FUNCTION "LKinCtrl_CallMC_Reset_SyncAxis" : Void   // FC35024, SCL
{ S7_Optimized_Access := 'TRUE' }
VERSION : 0.1
   VAR_INPUT
      syncAxisIn : TO_SynchronousAxis;   // SynchronousAxis to access
      execute : Bool;   // execute signal for MC_RESET
      restart : Bool;   // restart signal for MC_RESET
   END_VAR
   VAR_IN_OUT
      instMC_Reset : MC_RESET;   // multi instance of MC_RESET
   END_VAR
BEGIN
   //================================================================================
   // SIEMENS AG
   // (c)Copyright 2019 All Rights Reserved
   //--------------------------------------------------------------------------------
   // Library: LKinCtrl
   // Tested with: S7-1517T-3 PN
   // Engineering: TIA Portal V15
   // Restrictions: -
   // Requirements: S7-1500T FW 2.5
   // Functionality: Call MC_Home
   // Support: tech.team.motioncontrol@siemens.com
   // Note: Parameter comments are only available in language 'English (United States)'
   //-----------------------------------------------------------------------------
   // Change log table:
   // Version    Date          Expert in charge    Changes applied
   // 01.00.00   27.02.2019    JR                  First released version
   //===========================================================================================

   // call MC_Reset
   #instMC_Reset(Axis:=#syncAxisIn,
                 Execute:=#execute,
                 Restart:=#restart);
END_FUNCTION

FUNCTION "LKinCtrl_CallMC_Reset_PosAxis" : Void   // FC35025, SCL
{ S7_Optimized_Access := 'TRUE' }
VERSION : 0.1
   VAR_INPUT
      posAxisIn : TO_PositioningAxis;   // PositioningAxis to access
      execute : Bool;   // execute signal for MC_RESET
      restart : Bool;   // restart signal for MC_RESET
   END_VAR
   VAR_IN_OUT
      instMC_Reset : MC_RESET;   // multi instance of MC_RESET
   END_VAR
BEGIN
   //================================================================================
   // SIEMENS AG
   // (c)Copyright 2019 All Rights Reserved
   //--------------------------------------------------------------------------------
   // Library: LKinCtrl
   // Tested with: S7-1517T-3 PN
   // Engineering: TIA Portal V15
   // Restrictions: -
   // Requirements: S7-1500T FW 2.5
   // Functionality: Call MC_Reset
   // Support: tech.team.motioncontrol@siemens.com
   // Note: Parameter comments are only available in language 'English (United States)'
   //-----------------------------------------------------------------------------
   // Change log table:
   // Version    Date          Expert in charge    Changes applied
   // 01.00.00   27.02.2019    JR                  First released version
   //===========================================================================================

   // call MC_Reset
   #instMC_Reset(Axis:=#posAxisIn,
                 Execute:=#execute,
                 Restart:=#restart);
END_FUNCTION

FUNCTION "LKinCtrl_CallMC_Home_SyncAxis" : Void   // FC35026, SCL
{ S7_Optimized_Access := 'TRUE' }
VERSION : 0.1
   VAR_INPUT
      syncAxisIn : TO_SynchronousAxis;   // SynchronousAxis to access
      execute : Bool;   // execute trigger
      position : LReal;   // home position
      mode : Int;   // homing mode
   END_VAR
   VAR_IN_OUT
      instMC_Home : MC_HOME;   // multi instance MC_HOME
   END_VAR
BEGIN
   //================================================================================
   // SIEMENS AG
   // (c)Copyright 2019 All Rights Reserved
   //--------------------------------------------------------------------------------
   // Library: LKinCtrl
   // Tested with: S7-1517T-3 PN
   // Engineering: TIA Portal V15
   // Restrictions: -
   // Requirements: S7-1500T FW 2.5
   // Functionality: Call MC_Home
   // Support: tech.team.motioncontrol@siemens.com
   // Note: Parameter comments are only available in language 'English (United States)'
   //-----------------------------------------------------------------------------
   // Change log table:
   // Version    Date          Expert in charge    Changes applied
   // 01.00.00   27.02.2019    JR                  First released version
   //===========================================================================================

   // call MC_Home
   #instMC_Home(Axis:=#syncAxisIn,
                Execute:=#execute,
                Position:=#position,
                Mode:=#mode);
END_FUNCTION

FUNCTION "LKinCtrl_CallMC_Power_PosAxis" : Void   // FC35027, SCL
{ S7_Optimized_Access := 'TRUE' }
VERSION : 0.1
   VAR_INPUT
      posAxisIn : TO_PositioningAxis;   // PositioningAxis to access
      enable : Bool;   // execute signal for MC_RESET
      startMode : DInt;   // startMode of axis
      stopMode : Int;   // stopMode of axis
   END_VAR
   VAR_IN_OUT
      instMC_Power : MC_POWER;   // multi instance of MC_RESET
   END_VAR
BEGIN
   //================================================================================
   // SIEMENS AG
   // (c)Copyright 2019 All Rights Reserved
   //--------------------------------------------------------------------------------
   // Library: LKinCtrl
   // Tested with: S7-1517T-3 PN
   // Engineering: TIA Portal V15
   // Restrictions: -
   // Requirements: S7-1500T FW 2.5
   // Functionality: Call MC_Power
   // Support: tech.team.motioncontrol@siemens.com
   // Note: Parameter comments are only available in language 'English (United States)'
   //-----------------------------------------------------------------------------
   // Change log table:
   // Version    Date          Expert in charge    Changes applied
   // 01.00.00   04.03.2019    JR                  First released version
   //===========================================================================================

   // call MC_Reset
   #instMC_Power(Axis:=#posAxisIn,
                 Enable:=#enable,
                 StartMode:=#startMode,
                 StopMode:=#stopMode);
END_FUNCTION

FUNCTION "LKinCtrl_CallMC_Power_SyncAxis" : Void   // FC35028, SCL
{ S7_Optimized_Access := 'TRUE' }
VERSION : 0.1
   VAR_INPUT
      syncAxisIn : TO_SynchronousAxis;   // SynchronousAxis to access
      enable : Bool;   // execute signal for MC_RESET
      startMode : DInt;   // startMode of axis
      stopMode : Int;   // stopMode of axis
   END_VAR
   VAR_IN_OUT
      instMC_Power : MC_POWER;   // multi instance of MC_RESET
   END_VAR
BEGIN
   //================================================================================
   // SIEMENS AG
   // (c)Copyright 2019 All Rights Reserved
   //--------------------------------------------------------------------------------
   // Library: LKinCtrl
   // Tested with: S7-1517T-3 PN
   // Engineering: TIA Portal V15
   // Restrictions: -
   // Requirements: S7-1500T FW 2.5
   // Functionality: Call MC_Power
   // Support: tech.team.motioncontrol@siemens.com
   // Note: Parameter comments are only available in language 'English (United States)'
   //-----------------------------------------------------------------------------
   // Change log table:
   // Version    Date          Expert in charge    Changes applied
   // 01.00.00   04.03.2019    JR                  First released version
   //===========================================================================================

   // call MC_Reset
   #instMC_Power(Axis:=#syncAxisIn,
                 Enable:=#enable,
                 StartMode:=#startMode,
                 StopMode:=#stopMode);
END_FUNCTION

// folder: LKinCtrl_Blocks/LKinCtrl_SubBlocks

FUNCTION_BLOCK "LKinCtrl_PreBuffer"   // FB35001, SCL
TITLE = LKinCtrl_PreBuffer
{ S7_Optimized_Access := 'TRUE' }
AUTHOR : tech.team.motioncontrol@siemens.com
FAMILY : LKinCtrl
VERSION : 2.4
// The FB is copying the commands of the user defined PathData structure to an internal structure to be used for parametrizing motion commands later.
   VAR_INPUT
      enable : Bool;   // TRUE: Enable functionality of FB
      initPathTransition : DInt := 0;   // parameter from MC_MovePath interface
      initBufferMode : DInt := 1;   // parameter from MC_MovePath interface
      initTransitionParameter : Array[1..5] of LReal;   // parameter from MC_MovePath interface
      initPos : Array[1..4] of LReal;   // initial position from TO_Kinematics
      OCSFrames : Array[1..3] of "LKinCtrl_typeFrame";   // OCS frames from TO_Kinematics
      configuration : "LKinCtrl_typeConfiguration";   // configuration structure
      to_Kinematics : TO_Kinematics;   // reference to the axesGroup
   END_VAR
   VAR_OUTPUT
      valid : Bool;   // TRUE: Valid set of output values available at the FB
      busy : Bool;   // TRUE: FB is not finished and new output values can be expected
      error : Bool;   // TRUE: An error occurred during the execution of the FB
      status : Word := 16#7000;   // 16#0000 - 16#7FFF: Status of the FB, 16#8000 - 16#FFFF: Error identification
      preBufferLockDueToConfigCmd : Bool;   // TRUE: lock of PreBuffer due to config command ==> no continue for MC execution, lock GET_CMD
      lastCmdIdPathData : DInt;   // last command ID found in PathData
      pathDataRetrievePointer : DInt;   // actual value of the retrieve pointer from PathData
   END_VAR
   VAR_IN_OUT
      preprocessingStop : Bool;   // preprocessing stop output to halt MC execution
      pathData : Variant;   // connected PathData
      pathDataPreBuf : "LKinCtrl_typePathData_PreBuf";   // pre buffered exertion of PathData to be executed
   END_VAR
   VAR
      statEnableOld : Bool;   // old value of 'enable' input for edge detection
      statValid : Bool;   // static value for output 'valid'
      statBusy : Bool;   // static value for output 'busy'
      statError : Bool;   // static value for output 'error'
      statErrorUserCleared : Bool;   // error occurred that can only be solved by user; rising edge at enable input necessary
      statErrorAutoCleared : Bool;   // error occurred that can be acknowledged by FB
      statStatus : Word := 16#7000;   // static value for output 'status'
      statStateMachine : DInt := 0;   // state in the state machine of the FB
      statDebugState : Bool;   // static variable to enable stepwise debugging of state machine
      statDisablingCompleted : Bool;   // TRUE: Disabling has been completed
      statAsynchAddPointerRestart : Bool;   // static storing information of overflow of pointer
      statNumberOfPathDataElements : Int;   // static storing PathData elements (counted internally)
      statNoRestarts : DInt;   // static storing count of restarts of pointer
      statPathDataType : USInt;   // static storing of PathData type (reduced/normal/advanced)
      statPathDataName : String["LKINCTRL_LENGTH_OF_PATHDATA_NAME"];   // static storing of PathData name
      statSubsequentDeactCmdCtr : Int;   // number of subsequent deactivated commands in PathData
      statCmdIsMotionCmd : Bool;   // static to signalize command is motion command
      statCoordSystemOld : DInt;   // static storing of the last coordinate system
      statLastCmdIdPathdata : DInt;   // static storing of the last cmd id in PathData
      statCmdAdded : Bool;   // static to signalize if at least one cmd was added to preBuffer
      statRetValCircModeConv : Word;   // return value of circMode conversion
      statRetValLastPos : Word;   // return value of last position calculation
      statLinkConstellation : DInt;   // static storing the link constellation
      statPathDataPointers : "LKinCtrl_typeAdvPointers";   // static storing of actual PathData pointers
      statPathDataCommand : "LKinCtrl_typePathDataElement";   // static storing of actual PathData command
      statParameterValid : Array[1.."LKINCTRL_NO_OF_VALID_BITS"] of Bool;   // static storing for parameter valid bits from pathData advanced
      statLastPos : Array[1..4] of LReal;   // static array storing lastPos of path motion
      statAuxPoint : Array[1..3] of LReal;   // static array storing lastAuxPoint of path motion
      statOffsetCompActivated : Bool;   // static storing if offset compensation is active
      statOffsetCompActivatedOld : Bool;   // static storing of last compensation active
      statOffsetCompFirstCmd : Bool;   // bit to signalize first cmd of offset compensation
      statToolLength : LReal;   // static storing for the tool length
      statToolRadius : LReal;   // static storing for the tool radius
      statPathPlane : Int;   // static storing for the working plane of the tool
      statCompDirection : Int;   // static storing for the compensation direction (left/right)
      statRetrievePointerIncCtr : DInt;   // counter to search in path data
      statSearchNBOAborted : Bool;   // static bit to signalize abortion of search
      statNBOLastPos : Array[1..4] of LReal;   // storage variable lastPos for offset compensation
      statPathCmdOffCompIn : "LKinCtrl_typeCOffPathDataIn";   // static storing for the source contour offset element
      statPathCmdOffCompOut : "LKinCtrl_typeCOffPathDataOut";   // static storing for the target contour offset element
      statRetValOffsetComp : "LKinCtrl_typeCOffReturn";   // return value of the offset calculation
      statPathCmdNBOCheck : "LKinCtrl_typePathDataElement";   // static for path command when searching NBO command
      statDebugMessage : String;   // debugging string for development only
      statDebugNextCmdFound : DInt;   // debug variable to show index of next command
      statDebugNextButOneCmdFound : DInt;   // debug variable to show index of next but one command
      instMC_KinematicsTransformation : MC_KINEMATICSTRANSFORMATION;   // multi instance FB MC_KinematicsTransformation
      instMC_InverseKinematicsTransformation : MC_INVERSEKINEMATICSTRANSFORMATION;   // multi instance FB MC_InverseKinematicsTransformation
   END_VAR
   VAR_TEMP
      tempEnable : Bool;   // Temporary value for input 'enable'
      tempCtr : Int;   // Temporary counter
      tempFlagCtr : Int;   // Temporary counter
      tempNBOCoordSystemOld : DInt;   // Temporary value for old coord system when searching NBO
      tempCmdLengthIsZero : Bool;   // Temporary return value
      tempValidNextCmdFound : Bool;   // Temporary return value
      tempValidNextButOneCmdFound : Bool;   // Temporary return value
      tempIndexOk : Bool;   // Temporary return value
      tempRetVal : Word;   // Temporary return value
      tempParameterValidNBO : Array[1.."LKINCTRL_NO_OF_VALID_BITS"] of Bool;   // static storing for parameter valid bits from pathData advanced
      tempPathData_advanced : REF_TO "LKinCtrl_typePathData_advanced";   // Reference to path data advanced
      tempPathData : REF_TO "LKinCtrl_typePathData";   // Reference to path data
      tempPathData_reduced : REF_TO "LKinCtrl_typePathData_reduced";   // Reference to path data reduced
   END_VAR
   VAR CONSTANT
      NO_PROCESSING : DInt := 0;   // FB_PreBuffer state machine constant
      GET_CMD : DInt := 20;   // FB_PreBuffer state machine constant
      REGULAR_CMD : DInt := 21;   // FB_PreBuffer state machine constant
      OFFSET_CALC : DInt := 22;   // FB_PreBuffer state machine constant
      CHECK_CMD : DInt := 23;   // FB_PreBuffer state machine constant
      CHECK_NEXT_CMD : DInt := 25;   // FB_PreBuffer state machine constant
      SEARCH_NBO : DInt := 26;   // FB_PreBuffer state machine constant
      PATHDATA_PREBUFFERED_COMPLETELY : DInt := 40;   // FB_PreBuffer state machine constant
      DISABLE_STATE : DInt := 100;   // FB state: Disabling
      STATUS_NO_ERROR_IN_COMMAND : Word := 16#0000;   // command parameters correct, no error
      STATUS_NO_CALL : Word := 16#7000;   // no job being currently processed
      STATUS_FIRST_CALL : Word := 16#7001;   // first call after incoming new job (rising edge 'execute')
      STATUS_SUBSEQUENT_CALL : Word := 16#7002;   // Subsequent call during active processing without further details
      STATUS_PATHDATA_PREBUF_FULL : Word := 16#7010;   // PathData_preBuffered full with new commands
      STATUS_ALL_CMDS_BUFFERED : Word := 16#7100;   // all cmds buffered into PathData_preBuffered
      ERR_UNDEFINED_STATE : Word := 16#8600;   // error due to an undefined state in state machine
      ERR_OFFSET_COMPENSATION : Word := 16#8261;   // error during offset calculation
      ERR_LASTPOS_CALCULATION : Word := 16#8262;   // error during calculation of previous target position
      ERR_INVALID_PATHDATA_TYPE : Word := 16#8263;   // error due to an unsupported pathdata type
   END_VAR
   // statParameterValid[4] := True;
   // statParameterValid[3] := True;
   // statParameterValid[2] := True;
   // statParameterValid[1] := True;
BEGIN
   //==========================================================================================
   // SIEMENS AG
   // (c)Copyright 2020 All Rights Reserved
   //------------------------------------------------------------------------------------------
   // Library: LKinCtrl
   // Tested with: S7-1517T-3 PN/DP
   // Engineering: TIA Portal V16
   // Restrictions: ---
   // Requirements: S7-1500T FW 2.8
   // Functionality: LKinCtrl_PreBuffer
   // The FB is copying the commands of the user defined PathData structure
   // to an internal structure (PathDataPreBuffered) to be used for parametrizing
   // the motion commands later. 
   // 
   // Support: tech.team.motioncontrol@siemens.com
   // Note: Parameter comments are only available in language 'English (United States)'
   //------------------------------------------------------------------------------------------
   // Change log table:
   // Version    Date          Expert in charge    Changes applied
   // 01.00.00   06.02.2018    JR                  First release version V1.0
   // 02.00.00   18.04.2019    JR / FR             V2.0
   // 02.01.00   28.05.2019    JR / FR             V2.1 for LKinLang
   // 02.01.01   03.07.2019    JR                  BugFix for circMode 3 in offset compensation
   // 02.01.02   08.07.2019    JR                  BugFix for contour offset parameterValid Bits (PreBuffer)
   // 02.01.03   15.07.2019    JR                  Fixes for Contour Offset & parameter valid bits (PreBuffer)
   // 02.01.04   09.08.2019    JR                  Removal of code duplicates by functions
   // 02.02.00   28.01.2020    JR / FR             V2.2: Added valueFlags and flagOnlyCmd 
   // 02.02.01   07.02.2020    FR / DF             V2.2.1: Reset retrieve pointer when PreBuffer is disabled
   // 02.03.00   14.04.2020    FR                  Added preprocessing stop for LKinLang; Partial FB rework; Added "OCSFrames" input
   // 02.03.01   16.07.2020    FR                  Initialize preprocessing stop
   // 02.04.00   04.08.2020    FR                  Added MoveDirect and ConveyorTracking
   //===========================================================================================

   #tempEnable := #enable; // Work with temporary value / create process image

   REGION ENABLING/DISABLING
       IF (#tempEnable = TRUE) AND (#statStatus = #STATUS_NO_CALL) THEN // Enable FB
           // First call; initialize FB
           #statValid := TRUE;
           #statBusy := TRUE;
           #statError := FALSE;
           #statErrorUserCleared := FALSE;
           #statErrorAutoCleared := FALSE;
           #statStatus := #STATUS_FIRST_CALL;

           // Initialize add pointer in PathData_PreBuffered is done in MovePath
           // #pathDataPreBuf.addPointer := 1;

           #statStateMachine := #GET_CMD; // State machine - start functionality

           // initialize functionality: reset of variables, diagnostics, etc.
           #statDisablingCompleted := FALSE;

           // Init bool to signlaize config cmd
           #statSearchNBOAborted := FALSE;
           #statCmdAdded := FALSE;

           // Initialize reload bit & variables
           #statAsynchAddPointerRestart := FALSE;
           #pathDataPreBuf.addPointerRestarted := FALSE;
           // initialize lastCmdId in PathData with non-reachable value
           #statLastCmdIdPathdata := -1;
           #statNoRestarts := 0;
           #statOffsetCompActivated := FALSE;
           #statSubsequentDeactCmdCtr := 0;
           #statRetValOffsetComp.returnValue := 16#0;
           #statRetValOffsetComp."region" := 0;
           #statRetValOffsetComp.subBlockNumber := 0;
           #statRetValOffsetComp.internalNumber := 0;

           // copy initial position as last position if coordinates are not programmed (parameter invalid)
           #statLastPos := #initPos;
           // Init last coord system to WCS
           #statCoordSystemOld := "CS_WCS";

           // Get initial link constellation
           #statLinkConstellation := DWORD_TO_DINT(#to_Kinematics.StatusKinematics.LinkConstellation);

           // Reset instances
           #instMC_InverseKinematicsTransformation(AxesGroup := #to_Kinematics,
                                                   Enable := FALSE);
           #instMC_KinematicsTransformation(AxesGroup := #to_Kinematics,
                                            Enable := FALSE);

           // Added FR 2019.03.27
           // PathData conversion (reduced, regular(no suffix), advanced)
           //===========================================================================================
           // Reset path data type
           #statPathDataType := 0;

           REGION PATHDATA_TYPE
               // Reduced PathData (no circular commands, no pointers)
               IF TypeOf(#pathData) = LKinCtrl_typePathData_reduced THEN
                   #tempPathData_reduced ?= #pathData;
                   #statPathDataType := "LKINCTRL_PATHDATA_TYPE_REDUCED";
                   // Get last cmdID & number of PathData elements
                   #statNumberOfPathDataElements := "LKINCTRL_NO_OF_PATHDATA_ELEMENTS_REDUCED";

                   // Initialize retrieve pointer in PathData (if no pointers available, only set local static pointer variable)
                   #statPathDataPointers.retrievePointer := 0;

                   // Regular PathData (no pointers)
               ELSIF TypeOf(#pathData) = LKinCtrl_typePathData THEN
                   #tempPathData ?= #pathData;
                   #statPathDataType := "LKINCTRL_PATHDATA_TYPE_NORMAL";
                   // Get last cmdID
                   #statNumberOfPathDataElements := "LKINCTRL_NO_OF_PATHDATA_ELEMENTS";

                   // Initialize retrieve pointer in PathData (if no pointers available, only set local static pointer variable)
                   #statPathDataPointers.retrievePointer := 0;

                   // Advanced PathData (all elements)
               ELSIF TypeOf(#pathData) = LKinCtrl_typePathData_advanced THEN
                   #tempPathData_advanced ?= #pathData;
                   #statPathDataType := "LKINCTRL_PATHDATA_TYPE_ADVANCED";
                   #statNumberOfPathDataElements := "LKINCTRL_NO_OF_PATHDATA_ELEMENTS_ADVANCED";

                   // Initialize retrieve pointer in PathData
                   #tempPathData_advanced<?OpDeref?>.pointers.retrievePointer := 0;
                   #statPathDataPointers := #tempPathData_advanced<?OpDeref?>.pointers;

               ELSE
                   // Error wrong path data type 
                   #statStatus := #ERR_INVALID_PATHDATA_TYPE;
                   #statErrorAutoCleared := TRUE;
                   // Set state machine to no processing
                   #statStateMachine := #NO_PROCESSING;
               END_IF;

               // Init preprocessing stop
               #preprocessingStop := #statPathDataPointers.preprocessingStop;

           END_REGION PATHDATA_TYPE


       ELSIF (#tempEnable = FALSE) AND (#statEnableOld = TRUE) THEN // Disable FB 
           #statStateMachine := #DISABLE_STATE;

       ELSIF (#statStatus = #STATUS_FIRST_CALL) THEN // Set status identifier of subsequent call
           #statStatus := #STATUS_SUBSEQUENT_CALL;
       END_IF;

       // Edge detection 'enable' input
       #statEnableOld := #tempEnable;

       // Save old variables
       IF #statOffsetCompActivatedOld = TRUE
           AND #statOffsetCompActivated = FALSE
       THEN
           #preBufferLockDueToConfigCmd := FALSE;
       END_IF;
       #statOffsetCompActivatedOld := #statOffsetCompActivated;
   END_REGION ENABLING/DISABLING


   IF (#statStatus = #STATUS_NO_CALL) THEN // Nothing to do -> End here to reduce "system load"
       RETURN;
   END_IF;

   REGION CYCLIC_INPUT

       // Added FR 2019.03.27: Renew pointers every cycle
       IF TypeOf(#pathData) = LKinCtrl_typePathData_reduced THEN
           #tempPathData_reduced ?= #pathData;
           #statPathDataType := "LKINCTRL_PATHDATA_TYPE_REDUCED";
       ELSIF TypeOf(#pathData) = LKinCtrl_typePathData THEN
           #tempPathData ?= #pathData;
           #statPathDataType := "LKINCTRL_PATHDATA_TYPE_NORMAL";
       ELSIF TypeOf(#pathData) = LKinCtrl_typePathData_advanced THEN
           #tempPathData_advanced ?= #pathData;
           #statPathDataType := "LKINCTRL_PATHDATA_TYPE_ADVANCED";

           // Reset stopre in pathdata
           IF #statPathDataPointers.preprocessingStop = TRUE AND #preprocessingStop = FALSE THEN
               #statPathDataPointers.preprocessingStop := FALSE;
               #tempPathData_advanced<?OpDeref?>.pointers.preprocessingStop := FALSE;
           END_IF;

           // Get pointers in every cycle
           #statPathDataPointers := #tempPathData_advanced<?OpDeref?>.pointers;
       ELSE
           // Error wrong path data type 
           #statStatus := #ERR_INVALID_PATHDATA_TYPE;
           #statErrorAutoCleared := TRUE;
           // Set state machine to no processing
           #statStateMachine := #NO_PROCESSING;
       END_IF;

   END_REGION CYCLIC_INPUT


   REGION STATE_MACHINE
       // STATE: FB_STATE_NO_PROCESSING
       // =======================================================================================================
       // FB_STATE_NO_PROCESSING: // No processing active (Note: this state must always be present and left empty)
       IF #statStateMachine = #NO_PROCESSING THEN
           // do nothing, wait here
           ;
       END_IF;


       REGION PATHDATA_PREBUFFERING
           // STATE: GET_CMD
           // =======================================================================================================  
           // GET_CMD: Get cmd from connected path data and copy to internal
           // Next state: CHECK_CMD
           IF #statStateMachine = #GET_CMD
               // AND #statDebugState = TRUE
           THEN
               REGION GET_CMD
                   // reset  variable for single step debugging of states
                   #statDebugState := FALSE;

                   // retrievePointer must not pass addPointer (no reading of empty slots), if addPointer was not restarted ==> retrievePointer may catch up, not pass
                   IF (#pathDataPreBuf.retrievePointer <= #pathDataPreBuf.addPointer AND #pathDataPreBuf.addPointerRestarted = FALSE
                       // avoid addPointer to restart in next cycle (addPointer at end of list) if retreivePointer is at 1st element of PathDataPreBuffered ==> ?!
                       AND NOT (#pathDataPreBuf.addPointer = "LKINCTRL_NO_OF_PATHDATA_PREBUFFER_ELEMENTS" AND #pathDataPreBuf.retrievePointer = 1))
                       // addPointer must not pass retrievePointer (no overwriting not read slots), if addPointer was restarted ==> addPointer may not catch up
                       OR (#pathDataPreBuf.addPointerRestarted = TRUE AND #pathDataPreBuf.retrievePointer > #pathDataPreBuf.addPointer + 1)
                       // add condition here to avoid addPointer catching up with retrievePointer after addPointerRestart (additional offset compensation command) 
                       // in case of intermediate command --> 2 commands get inserted --> additional buffer check is needed
                       // --> See release notes in OneNote
                       // add into brackets of OR statement above
                       // // AND NOT ()
                   THEN
                       // Path command copy procedure
                       //------------------------------------------------------------------------------------------
                       // INSERT PATH DATA RING BUFFER FUNCTIONALITY HERE
                       // ring buffer code => TO be tested
                       // Condition 1: ignore addPointer if no ring buffer is running (PathData_regular/PathData_reduced attached)
                       IF (#statPathDataPointers.ignoreAddPointer = TRUE)
                           // Condition 2: respect addPointer (PathData_advanced attached) - regular ring buffer limiatations 
                           OR
                           ((#statPathDataPointers.ignoreAddPointer = FALSE)
                           AND (#statPathDataPointers.bufferLocked = FALSE)
                           AND (
                           // retrievePointer must not pass addPointer (no reading of empty slots), if addPointer was not restarted ==> retrievePointer may catch up, not pass
                           // FR 26.04.2019: changed from <= to <
                           ((#statPathDataPointers.retrievePointer < #statPathDataPointers.addPointer AND #statPathDataPointers.addPointerRestarted = FALSE)
                           // addPointer must not pass retrievePointer (no overwriting not read slots), if addPointer was restarted ==> addPointer may not catch up
                           OR (#statPathDataPointers.retrievePointer > #statPathDataPointers.addPointer AND #statPathDataPointers.addPointerRestarted = TRUE))))
                       THEN

                           // increase PathData retreivePointer
                           IF #statPathDataPointers.retrievePointer <= #statNumberOfPathDataElements
                           THEN
                               #statPathDataPointers.retrievePointer += 1;
                           END_IF;

                           // Ring buffer
                           IF #statPathDataPointers.retrievePointer > #statNumberOfPathDataElements AND NOT #statPathDataPointers.ignoreAddPointer THEN
                               #statPathDataPointers.retrievePointer := 1;
                               // set addPointer restart bit
                               #statPathDataPointers.addPointerRestarted := FALSE;
                               // count restart cycles of PathData retrievePointer
                               #statNoRestarts += 1;
                           END_IF;

                           // check for length of PathData array to do not exceed element count
                           IF #statPathDataPointers.retrievePointer <= #statNumberOfPathDataElements
                               AND #statPathDataPointers.retrievePointer > 0
                           THEN

                               // Copy actual path data element where retrievePointer is pointing at
                               IF #statPathDataType = "LKINCTRL_PATHDATA_TYPE_REDUCED" THEN
                                   // Get name of path data
                                   #statPathDataName := #tempPathData_reduced<?OpDeref?>.pathDataName;
                               ELSIF #statPathDataType = "LKINCTRL_PATHDATA_TYPE_NORMAL" THEN
                                   // Get name of path data
                                   #statPathDataName := #tempPathData<?OpDeref?>.pathDataName;
                               ELSIF #statPathDataType = "LKINCTRL_PATHDATA_TYPE_ADVANCED" THEN
                                   // Get name of path data
                                   #statPathDataName := #tempPathData_advanced<?OpDeref?>.pathDataName;
                               ELSE
                                   // Error wrong path data type 
                                   #statStatus := #ERR_INVALID_PATHDATA_TYPE;
                                   #statErrorAutoCleared := TRUE;
                                   // Set state machine to no processing
                                   #statStateMachine := #NO_PROCESSING;
                               END_IF;

                               // Copy path command from path data
                               #tempRetVal := "LKinCtrl_GetPathDataCmd"(pathDataType := #statPathDataType,
                                                                        index := #statPathDataPointers.retrievePointer,
                                                                        pathDataReduced := #tempPathData_reduced,
                                                                        pathData := #tempPathData,
                                                                        pathDataAdvanced := #tempPathData_advanced,
                                                                        pathDataCommand => #statPathDataCommand,
                                                                        parameterValid => #statParameterValid);

                               // check for command to be deactivated
                               IF #statPathDataCommand.cmdActivated THEN
                                   // Go to check cmd state
                                   #statStateMachine := #CHECK_CMD;
                               ELSE
                                   // count subsequent deactivated commands
                                   #statSubsequentDeactCmdCtr += 1;
                                   // do nothing as pathData.retrievePointer has already been increased ==> next cmd checked in next cycle
                               END_IF;
                           ELSE
                               // end of PathData array reached ==> do nothing?
                               // set status to show pre buffering is completed ==> external disable in next state of MovePath
                               #statStatus := #STATUS_ALL_CMDS_BUFFERED;
                               // set stateMachine
                               #statStateMachine := #PATHDATA_PREBUFFERED_COMPLETELY;
                           END_IF;
                       END_IF;
                   ELSE
                       // PathDataPreBuf full
                       // FB has not transferred the next cmd to the addPointer element in PathDataPreBuf yet
                       // set status 
                       #statStatus := #STATUS_PATHDATA_PREBUF_FULL;
                   END_IF;
               END_REGION GET_CMD
           END_IF;

           // STATE: CHECK_CMD
           // =======================================================================================================   
           // CHECK_CMD: Check cmd if executable and if offset comp is activated
           IF #statStateMachine = #CHECK_CMD THEN
               REGION CHECK_CMD
                   // check for command to be last command (today also end of PathData: -1) 
                   IF #statPathDataCommand.cmdType < 0 THEN
                       // last activated command in PathData reached
                       // set status to show pre buffering is completed
                       #statStatus := #STATUS_ALL_CMDS_BUFFERED;
                       // set stateMachine
                       #statStateMachine := #PATHDATA_PREBUFFERED_COMPLETELY;
                   ELSE
                       // reset counter of subsequent deactivated commands when command is activated and not 'End of List'
                       #statSubsequentDeactCmdCtr := 0;

                       // command check in external FC
                       #statStatus := "LKinCtrl_CheckPathDataCmd"(cmdIsMotionCmd => #statCmdIsMotionCmd,
                                                                  pathDataCmd := #statPathDataCommand);

                       // Check for moveDirect command during ContourOffset
                       IF #statStatus = #STATUS_NO_ERROR_IN_COMMAND
                           AND #statOffsetCompActivated = TRUE
                           AND (#statPathDataCommand.cmdType = "LKINCTRL_MC_MOVEDIRECTABS"
                           OR #statPathDataCommand.cmdType = "LKINCTRL_MC_MOVEDIRECTREL")
                       THEN
                           // Set error status 
                           #statStatus := #ERR_OFFSET_COMPENSATION;
                       END_IF;

                       // check if no error was detected ==> command configured correctly
                       IF #statStatus = #STATUS_NO_ERROR_IN_COMMAND THEN

                           // PathData - general - information
                           //====================================================================================================================================
                           #pathDataPreBuf.commands[#pathDataPreBuf.addPointer].pathDataName := #statPathDataName;

                           // command is no intermediate command by default, only changed with actived offset compensation and generation of additional command
                           #pathDataPreBuf.commands[#pathDataPreBuf.addPointer].isIntermediateCmd := FALSE;

                           // PathData command 
                           //====================================================================================================================================
                           //PathData - command - cmdType
                           IF #statPathDataCommand.cmdType = "LKINCTRL_CONFIG_START_OFFSET_COMP_LEFT"      // configuration command - offset compensation activated left
                               OR #statPathDataCommand.cmdType = "LKINCTRL_CONFIG_START_OFFSET_COMP_RIGHT"   // configuration command - offset compensation activated right
                           THEN
                               // handle activation of contour offset calculation
                               #statOffsetCompActivated := TRUE;
                               #statOffsetCompFirstCmd := TRUE;
                               #preBufferLockDueToConfigCmd := TRUE;

                               // store compensation calculation parameters
                               #statToolLength := #configuration.offsetParameter[#statPathDataCommand.cmdParameters.offsetParameters.offsetParaNo].length;
                               #statToolRadius := #configuration.offsetParameter[#statPathDataCommand.cmdParameters.offsetParameters.offsetParaNo].radius;
                               #statPathPlane := #statPathDataCommand.cmdParameters.offsetParameters.mainPathPlane;

                               // If lastPos is in MCS then transform to WCS as Contour offset needs cartesian coordinates!
                               IF #statCoordSystemOld = "CS_MCS" THEN
                                   // Transform lastPos to WCS
                                   #instMC_KinematicsTransformation(AxesGroup := #to_Kinematics,
                                                                    Enable := TRUE,
                                                                    AxesPosition := #statLastPos,
                                                                    CoordSystem := "CS_WCS",
                                                                    ErrorId=>#tempRetVal,
                                                                    Position => #statLastPos,
                                                                    LinkConstellation => #statLinkConstellation);

                                   // Update old coordSystem
                                   #statCoordSystemOld := "CS_WCS";

                                   // check for error in last position calculation
                                   IF #tempRetVal <> 16#0 THEN
                                       // set error status
                                       #statErrorAutoCleared := TRUE;
                                       #statStatus := #tempRetVal;
                                   END_IF;
                               END_IF;

                               // Initial position
                               #statPathCmdOffCompIn.currentPos.positionAbsolute.x := #statLastPos[1];
                               #statPathCmdOffCompIn.currentPos.positionAbsolute.y := #statLastPos[2];
                               #statPathCmdOffCompIn.currentPos.positionAbsolute.z := #statLastPos[3];
                               #statPathCmdOffCompIn.currentPos.positionAbsolute.a := #statLastPos[4];

                               // added according to AW
                               #statPathCmdOffCompIn.currentPos.positionAbsoluteRadComp := #statPathCmdOffCompIn.currentPos.positionAbsolute;

                               IF #statPathDataCommand.cmdType = "LKINCTRL_CONFIG_START_OFFSET_COMP_LEFT" THEN
                                   // store compensation calculation parameters
                                   #statCompDirection := "LKINCTRL_COMP_LEFT";

                               ELSIF #statPathDataCommand.cmdType = "LKINCTRL_CONFIG_START_OFFSET_COMP_RIGHT" THEN
                                   // store compensation calculation parameters
                                   #statCompDirection := "LKINCTRL_COMP_RIGHT";
                               END_IF;

                               // Go to copy cmd
                               #statStateMachine := #GET_CMD;

                           ELSIF #statPathDataCommand.cmdType = "LKINCTRL_CONFIG_END_OFFSET_COMP" THEN       // configuration command - offset compensation deactivated
                               IF #statOffsetCompActivated THEN // Only do this if the offset comp was actually activated
                                   // handle deactivation of contour offset calculation
                                   #statOffsetCompActivated := FALSE;

                                   // update last pos when deactivating contour offset
                                   // --> Keep corrected positions as "modal"
                                   #statLastPos[1] := #statPathCmdOffCompOut.nextPositionAbsoluteRadComp.x;
                                   #statLastPos[2] := #statPathCmdOffCompOut.nextPositionAbsoluteRadComp.y;
                                   #statLastPos[3] := #statPathCmdOffCompOut.nextPositionAbsoluteRadComp.z;
                                   #statLastPos[4] := #statPathCmdOffCompOut.nextPositionAbsoluteRadComp.a;
                               END_IF;

                               // Go to copy cmd
                               #statStateMachine := #GET_CMD;

                           ELSE // regular motion command

                               // Set bit to signal at least one cmd is added to preBuffered
                               #statCmdAdded := TRUE;

                               // handle regular command copying
                               IF #statOffsetCompActivated = FALSE OR #statCmdIsMotionCmd = FALSE THEN
                                   #statStateMachine := #REGULAR_CMD;
                               ELSE // Compensation active
                                   #statStateMachine := #CHECK_NEXT_CMD;
                               END_IF;

                           END_IF;
                       ELSE
                           // Error in command 
                           #statErrorAutoCleared := TRUE;
                       END_IF;
                   END_IF;
               END_REGION CHECK_CMD
           END_IF;

           // STATE: REGULAR_CMD
           // =======================================================================================================   
           // REGULAR_CMD: Copy regular cmd
           IF #statStateMachine = #REGULAR_CMD THEN
               REGION COPY_CMD_REGULAR
                   //PathData - command - cmdType
                   #pathDataPreBuf.commands[#pathDataPreBuf.addPointer].cmdType := #statPathDataCommand.cmdType;

                   //PathData - command - cmdID
                   #pathDataPreBuf.commands[#pathDataPreBuf.addPointer].cmdID := #statPathDataPointers.retrievePointer + #statNoRestarts * INT_TO_DINT("LKINCTRL_NO_OF_PATHDATA_ELEMENTS_ADVANCED");

                   //PathData - command - cmdName
                   #pathDataPreBuf.commands[#pathDataPreBuf.addPointer].cmdName := #statPathDataCommand.cmdName;

                   // Copy validBits to PreBuffer 03.05.2019 FR
                   // PathData - command - ValidBits
                   #pathDataPreBuf.commands[#pathDataPreBuf.addPointer].parameterValid := #statParameterValid;

                   //PathData - command - cmdCoordinates
                   //====================================================================================================================================
                   //PathData - command - cmdCoordinates - absolutePosition[1..4]
                   #pathDataPreBuf.commands[#pathDataPreBuf.addPointer].cmdCoordinates.absolutePosition[1] := #statPathDataCommand.cmdCoordinates.cartesianPosition.x;
                   #pathDataPreBuf.commands[#pathDataPreBuf.addPointer].cmdCoordinates.absolutePosition[2] := #statPathDataCommand.cmdCoordinates.cartesianPosition.y;
                   #pathDataPreBuf.commands[#pathDataPreBuf.addPointer].cmdCoordinates.absolutePosition[3] := #statPathDataCommand.cmdCoordinates.cartesianPosition.z;
                   #pathDataPreBuf.commands[#pathDataPreBuf.addPointer].cmdCoordinates.absolutePosition[4] := #statPathDataCommand.cmdCoordinates.cartesianPosition.a;

                   //PathData - command - cmdCoordinates - coordSystem
                   #pathDataPreBuf.commands[#pathDataPreBuf.addPointer].cmdCoordinates.coordSystem := #statPathDataCommand.cmdCoordinates.coordSystem;


                   //PathData - command - cmdParameters
                   //====================================================================================================================================
                   #pathDataPreBuf.commands[#pathDataPreBuf.addPointer].cmdParameters := #statPathDataCommand.cmdParameters;


                   //PathData - command - setFlags
                   //====================================================================================================================================
                   // also copy flagMode to pathDataPreBuf for use in specific case of waitFlag
                   FOR #tempFlagCtr := 1 TO "LKINCTRL_NO_OF_CMD_SETFLAGS" DO
                       #pathDataPreBuf.commands[#pathDataPreBuf.addPointer].setFlags[#tempFlagCtr] := #statPathDataCommand.setFlags[#tempFlagCtr];
                       // // change flagMode 3 to flagMode 2 as functionality is equal
                       // check for cmd to be flagOnly cmd
                       // check for cmd to implement flag and flagMode to be flagMode 3
                       IF #pathDataPreBuf.commands[#pathDataPreBuf.addPointer].cmdType = "LKINCTRL_CMD_FLAG_ONLY"
                           AND #pathDataPreBuf.commands[#pathDataPreBuf.addPointer].setFlags[#tempFlagCtr].flag <> -1
                           AND #pathDataPreBuf.commands[#pathDataPreBuf.addPointer].setFlags[#tempFlagCtr].flagMode = 3
                       THEN
                           // change flagMode 3 to flagMode 2
                           #pathDataPreBuf.commands[#pathDataPreBuf.addPointer].setFlags[#tempFlagCtr].flagMode := 2;
                       END_IF;
                   END_FOR;